HMI tags "Robot"
   "name" : Int, internal
   "DB1901_Config_Robots_Config_Robots{0}_Type_Kuka" : Bool = PLC DB1901_Config_Robots.Config_Robots[0].Type_Kuka AT %DB1901.DBX6.0, 1 s
      on ChangeValue: SetBit("DB1901_Config_Robots_Write")
   "DB1901_Config_Robots_Config_Robots{0}_Type_ABB" : Bool = PLC DB1901_Config_Robots.Config_Robots[0].Type_ABB AT %DB1901.DBX6.1, 1 s
      on ChangeValue: SetBit("DB1901_Config_Robots_Write")
   "DB1901_Config_Robots_Config_Robots{0}_Type_Fanuc" : Bool = PLC DB1901_Config_Robots.Config_Robots[0].Type_Fanuc AT %DB1901.DBX6.2, 1 s
      on ChangeValue: SetBit("DB1901_Config_Robots_Write")
   "DB1901_Config_Robots_Config_Robots{0}_Type_Motoman" : Bool = PLC DB1901_Config_Robots.Config_Robots[0].Type_Motoman AT %DB1901.DBX6.3, 1 s
      on ChangeValue: SetBit("DB1901_Config_Robots_Write")
   "DB1901_Config_Robots_Config_Robots{0}_Type_5" : Bool = PLC DB1901_Config_Robots.Config_Robots[0].Type_5 AT %DB1901.DBX6.4, 1 s
      on ChangeValue: SetBit("DB1901_Config_Robots_Write")
   "DB1901_Config_Robots_Config_Robots{0}_Type_6" : Bool = PLC DB1901_Config_Robots.Config_Robots[0].Type_6 AT %DB1901.DBX6.5, 1 s
      on ChangeValue: SetBit("DB1901_Config_Robots_Write")
   "DB1901_Config_Robots_Config_Robots{0}_Type_7" : Bool = PLC DB1901_Config_Robots.Config_Robots[0].Type_7 AT %DB1901.DBX6.6, 1 s
      on ChangeValue: SetBit("DB1901_Config_Robots_Write")
   "DB1901_Config_Robots_Config_Robots{0}_Type_8" : Bool = PLC DB1901_Config_Robots.Config_Robots[0].Type_8 AT %DB1901.DBX6.7, 1 s
      on ChangeValue: SetBit("DB1901_Config_Robots_Write")
   "DB1901_Config_Robots_Config_Robots{0}_With_Shotware" : Bool = PLC DB1901_Config_Robots.Config_Robots[0].With_Shotware AT %DB1901.DBX7.0, 1 s
      on ChangeValue: SetBit("DB1901_Config_Robots_Write")
   "DB1901_Config_Robots_Config_Robots{0}_With_Tracking" : Bool = PLC DB1901_Config_Robots.Config_Robots[0].With_Tracking AT %DB1901.DBX7.1, 1 s
      on ChangeValue: SetBit("DB1901_Config_Robots_Write")
   "DB1901_Config_Robots_Config_Robots{0}_With_Safetysoftware" : Bool = PLC DB1901_Config_Robots.Config_Robots[0].With_Safetysoftware AT %DB1901.DBX7.2, 1 s
      on ChangeValue: SetBit("DB1901_Config_Robots_Write")
   "DB1901_Config_Robots_Config_Robots{0}_With_Synchronisation" : Bool = PLC DB1901_Config_Robots.Config_Robots[0].With_Synchronisation AT %DB1901.DBX7.3, 1 s
      on ChangeValue: SetBit("DB1901_Config_Robots_Write")
   "DB1901_Config_Robots_Config_Robots{0}_With_Testshot" : Bool = PLC DB1901_Config_Robots.Config_Robots[0].With_Testshot AT %DB1901.DBX7.4, 1 s
      on ChangeValue: SetBit("DB1901_Config_Robots_Write")
   "DB1901_Config_Robots_Config_Robots{0}_With_Cleaning" : Bool = PLC DB1901_Config_Robots.Config_Robots[0].With_Cleaning AT %DB1901.DBX7.5, 1 s
      on ChangeValue: SetBit("DB1901_Config_Robots_Write")
   "DB1901_Config_Robots_Config_Robots{0}_With_Wet_Cleaning" : Bool = PLC DB1901_Config_Robots.Config_Robots[0].With_Wet_Cleaning AT %DB1901.DBX7.6, 1 s
      on ChangeValue: SetBit("DB1901_Config_Robots_Write")
   "DB1901_Config_Robots_Config_Robots{0}_With_Wet_Cleaning_LFI" : Bool = PLC DB1901_Config_Robots.Config_Robots[0].With_Wet_Cleaning_LFI AT %DB1901.DBX7.7, 1 s
      on ChangeValue: SetBit("DB1901_Config_Robots_Write")
   "DB1901_Config_Robots_Config_Robots{0}_With_Wet_Cleaning_Spray" : Bool = PLC DB1901_Config_Robots.Config_Robots[0].With_Wet_Cleaning_Spray AT %DB1901.DBX8.0, 1 s
      on ChangeValue: SetBit("DB1901_Config_Robots_Write")
   "DB1901_Config_Robots_Config_Robots{0}_With_IR_Station" : Bool = PLC DB1901_Config_Robots.Config_Robots[0].With_IR_Station AT %DB1901.DBX8.1, 1 s
      on ChangeValue: SetBit("DB1901_Config_Robots_Write")
   "DB1901_Config_Robots_Config_Robots{0}_With_Brush_Station" : Bool = PLC DB1901_Config_Robots.Config_Robots[0].With_Brush_Station AT %DB1901.DBX8.2, 1 s
      on ChangeValue: SetBit("DB1901_Config_Robots_Write")
   "DB1901_Config_Robots_Config_Robots{0}_With_Belt_Filter" : Bool = PLC DB1901_Config_Robots.Config_Robots[0].With_Belt_Filter AT %DB1901.DBX8.3, 1 s
      on ChangeValue: SetBit("DB1901_Config_Robots_Write")
   "DB1901_Config_Robots_Config_Robots{0}_With_Air_Cleaner" : Bool = PLC DB1901_Config_Robots.Config_Robots[0].With_Air_Cleaner AT %DB1901.DBX8.4, 1 s
      on ChangeValue: SetBit("DB1901_Config_Robots_Write")
   "DB1901_Config_Robots_Config_Robots{0}_Spare_2_5" : Bool = PLC DB1901_Config_Robots.Config_Robots[0].Spare_2_5 AT %DB1901.DBX8.5, 1 s
      on ChangeValue: SetBit("DB1901_Config_Robots_Write")
   "DB1901_Config_Robots_Config_Robots{0}_Spare_2_6" : Bool = PLC DB1901_Config_Robots.Config_Robots[0].Spare_2_6 AT %DB1901.DBX8.6, 1 s
      on ChangeValue: SetBit("DB1901_Config_Robots_Write")
   "DB1901_Config_Robots_Config_Robots{0}_Spare_2_7" : Bool = PLC DB1901_Config_Robots.Config_Robots[0].Spare_2_7 AT %DB1901.DBX8.7, 1 s
      on ChangeValue: SetBit("DB1901_Config_Robots_Write")
   "DB1900_IF_Robots_State_Robots{0}_EmergencyStopReady" : Bool = PLC DB1900_IF_Robots.State_Robots[0].EmergencyStopReady AT %DB1900.DBX96.4, 1 s
   "DB1900_IF_Robots_State_Robots{0}_AutomatcStopReady" : Bool = PLC DB1900_IF_Robots.State_Robots[0].AutomatcStopReady AT %DB1900.DBX96.5, 1 s
   "DB1900_IF_Robots_State_Robots{0}_MixingheadAuto" : Bool = PLC DB1900_IF_Robots.State_Robots[0].MixingheadAuto AT %DB1900.DBX96.6, 1 s
   "DB1900_IF_Robots_State_Robots{0}_MaschineAuto" : Bool = PLC DB1900_IF_Robots.State_Robots[0].MaschineAuto AT %DB1900.DBX96.7, 1 s
   "DB1900_IF_Robots_State_Robots{0}_TestShotRunning" : Bool = PLC DB1900_IF_Robots.State_Robots[0].TestShotRunning AT %DB1900.DBX97.3, 1 s
   "DB1900_IF_Robots_State_Robots{0}_Rob_in_Home" : Bool = PLC DB1900_IF_Robots.State_Robots[0].Rob_in_Home AT %DB1900.DBX96.0, 1 s
   "DB1900_IF_Robots_State_Robots{0}_Rob_in_Automatic" : Bool = PLC DB1900_IF_Robots.State_Robots[0].Rob_in_Automatic AT %DB1900.DBX96.1, 1 s
   "DB1900_IF_Robots_State_Robots{0}_Rob_in_Cycle" : Bool = PLC DB1900_IF_Robots.State_Robots[0].Rob_in_Cycle AT %DB1900.DBX96.2, 1 s
   "DB1900_IF_Robots_Switch_Robots{0}_SwitchHomePosON_OFF" : Bool = PLC DB1900_IF_Robots.Switch_Robots[0].SwitchHomePosON_OFF AT %DB1900.DBX6.0, 1 s
      on ChangeValue: SetBit("DB1900_IF_Robots_Write")
   "DB1900_IF_Robots_Switch_Robots{0}_SwitchMaintPosON_OFF" : Bool = PLC DB1900_IF_Robots.Switch_Robots[0].SwitchMaintPosON_OFF AT %DB1900.DBX6.1, 1 s
      on ChangeValue: SetBit("DB1900_IF_Robots_Write")
   "DB1900_IF_Robots_Switch_Robots{0}_SwitchMaintPos_2ON_OFF" : Bool = PLC DB1900_IF_Robots.Switch_Robots[0].SwitchMaintPos_2ON_OFF AT %DB1900.DBX6.2, 1 s
      on ChangeValue: SetBit("DB1900_IF_Robots_Write")
   "DB1900_IF_Robots_Switch_Robots{0}_SwitchTestShotON_OFF" : Bool = PLC DB1900_IF_Robots.Switch_Robots[0].SwitchTestShotON_OFF AT %DB1900.DBX6.3, 1 s
      on ChangeValue: SetBit("DB1900_IF_Robots_Write")
   "DB1900_IF_Robots_Switch_Robots{0}_SwitchCleaningON_OFF" : Bool = PLC DB1900_IF_Robots.Switch_Robots[0].SwitchCleaningON_OFF AT %DB1900.DBX6.4, 1 s
      on ChangeValue: SetBit("DB1900_IF_Robots_Write")
   "DB1900_IF_Robots_Switch_Robots{0}_SwitchBrushON_OFF" : Bool = PLC DB1900_IF_Robots.Switch_Robots[0].SwitchBrushON_OFF AT %DB1900.DBX6.5, 1 s
      on ChangeValue: SetBit("DB1900_IF_Robots_Write")
   "DB1900_IF_Robots_Switch_Robots{0}_SwitchSyncON_OFF" : Bool = PLC DB1900_IF_Robots.Switch_Robots[0].SwitchSyncON_OFF AT %DB1900.DBX6.6, 1 s
      on ChangeValue: SetBit("DB1900_IF_Robots_Write")
   "DB1900_IF_Robots_Switch_Robots{0}_SwitchTeachenON_OFF" : Bool = PLC DB1900_IF_Robots.Switch_Robots[0].SwitchTeachenON_OFF AT %DB1900.DBX6.7, 1 s
      on ChangeValue: SetBit("DB1900_IF_Robots_Write")
   "DB1900_IF_Robots_Switch_Robots{0}_SwitchLearningON_OFF" : Bool = PLC DB1900_IF_Robots.Switch_Robots[0].SwitchLearningON_OFF AT %DB1900.DBX7.0, 1 s
      on ChangeValue: SetBit("DB1900_IF_Robots_Write")
   "DB1900_IF_Robots_Switch_Robots{0}_SwitchAirCleaningON_OFF" : Bool = PLC DB1900_IF_Robots.Switch_Robots[0].SwitchAirCleaningON_OFF AT %DB1900.DBX7.1, 1 s
      on ChangeValue: SetBit("DB1900_IF_Robots_Write")
   "DB1900_IF_Robots_Switch_Robots{0}_SwitchAirCleaningManON_OFF" : Bool = PLC DB1900_IF_Robots.Switch_Robots[0].SwitchAirCleaningManON_OFF AT %DB1900.DBX7.2, 1 s
      on ChangeValue: SetBit("DB1900_IF_Robots_Write")
   "DB1900_IF_Robots_Switch_Robots{0}_StateHomePos" : Byte = PLC DB1900_IF_Robots.Switch_Robots[0].StateHomePos AT %DB1900.DBB8, 1 s
      on ChangeValue: SetBit("DB1900_IF_Robots_Write")
   "DB1900_IF_Robots_Switch_Robots{0}_StateMaintPos" : Byte = PLC DB1900_IF_Robots.Switch_Robots[0].StateMaintPos AT %DB1900.DBB9, 1 s
      on ChangeValue: SetBit("DB1900_IF_Robots_Write")
   "DB1900_IF_Robots_Switch_Robots{0}_StateMaintPos_2" : Byte = PLC DB1900_IF_Robots.Switch_Robots[0].StateMaintPos_2 AT %DB1900.DBB10, 1 s
      on ChangeValue: SetBit("DB1900_IF_Robots_Write")
   "DB1900_IF_Robots_Switch_Robots{0}_StateTestShot" : Byte = PLC DB1900_IF_Robots.Switch_Robots[0].StateTestShot AT %DB1900.DBB11, 1 s
      on ChangeValue: SetBit("DB1900_IF_Robots_Write")
   "DB1900_IF_Robots_Switch_Robots{0}_StateCleaning" : Byte = PLC DB1900_IF_Robots.Switch_Robots[0].StateCleaning AT %DB1900.DBB12, 1 s
      on ChangeValue: SetBit("DB1900_IF_Robots_Write")
   "DB1900_IF_Robots_Switch_Robots{0}_StateBrush" : Byte = PLC DB1900_IF_Robots.Switch_Robots[0].StateBrush AT %DB1900.DBB13, 1 s
      on ChangeValue: SetBit("DB1900_IF_Robots_Write")
   "DB1900_IF_Robots_Switch_Robots{0}_StateSync" : Byte = PLC DB1900_IF_Robots.Switch_Robots[0].StateSync AT %DB1900.DBB14, 1 s
      on ChangeValue: SetBit("DB1900_IF_Robots_Write")
   "DB1900_IF_Robots_Switch_Robots{0}_StateTeachen" : Byte = PLC DB1900_IF_Robots.Switch_Robots[0].StateTeachen AT %DB1900.DBB15, 1 s
      on ChangeValue: SetBit("DB1900_IF_Robots_Write")
   "DB1900_IF_Robots_Switch_Robots{0}_StateLearning" : Byte = PLC DB1900_IF_Robots.Switch_Robots[0].StateLearning AT %DB1900.DBB16, 1 s
      on ChangeValue: SetBit("DB1900_IF_Robots_Write")
   "DB1900_IF_Robots_Switch_Robots{0}_StateAirCleaning" : Byte = PLC DB1900_IF_Robots.Switch_Robots[0].StateAirCleaning AT %DB1900.DBB17, 1 s
      on ChangeValue: SetBit("DB1900_IF_Robots_Write")
   "DB1900_IF_Robots_Switch_Robots{0}_StateAirCleaningManual" : Byte = PLC DB1900_IF_Robots.Switch_Robots[0].StateAirCleaningManual AT %DB1900.DBB18, 1 s
      on ChangeValue: SetBit("DB1900_IF_Robots_Write")
   "DB1900_IF_Robots_ReadWriteDeviceNo" : Int = PLC DB1900_IF_Robots.ReadWriteDeviceNo AT %DB1900.DBW0, 1 s
   "DB1900_IF_Robots_Read" : Bool = PLC DB1900_IF_Robots.Read AT %DB1900.DBX4.0, 1 s
   "DB1900_IF_Robots_Write" : Bool = PLC DB1900_IF_Robots.Write AT %DB1900.DBX4.1, 1 s
   "DB1901_Config_Robots_Read" : Bool = PLC DB1901_Config_Robots.Read AT %DB1901.DBX4.0, 1 s
   "DB1901_Config_Robots_Write" : Bool = PLC DB1901_Config_Robots.Write AT %DB1901.DBX4.1, 1 s
   "DB1900_IF_Robots_State_Robots{0}_Rob_Prog_No" : Byte = PLC DB1900_IF_Robots.State_Robots[0].Rob_Prog_No AT %DB1900.DBB98, 1 s
   "DB1900_IF_Robots_State_Robots{0}_Rob_MC_No" : Byte = PLC DB1900_IF_Robots.State_Robots[0].Rob_MC_No AT %DB1900.DBB99, 1 s

HMI tags "Navigation Button"
   "DB14_TP_Shortcuts_TP_Shortcuts_ButtonNo_1" : Bool = PLC DB14_TP_Shortcuts.TP_Shortcuts.ButtonNo.1, 1 s
   "DB14_TP_Shortcuts_TP_Shortcuts_ButtonNo_2" : Bool = PLC DB14_TP_Shortcuts.TP_Shortcuts.ButtonNo.2, 1 s
   "DB14_TP_Shortcuts_TP_Shortcuts_ButtonNo_3" : Bool = PLC DB14_TP_Shortcuts.TP_Shortcuts.ButtonNo.3, 1 s
   "DB14_TP_Shortcuts_TP_Shortcuts_ButtonNo_5" : Bool = PLC DB14_TP_Shortcuts.TP_Shortcuts.ButtonNo.5, 1 s
   "DB14_TP_Shortcuts_TP_Shortcuts_ButtonNo_6" : Bool = PLC DB14_TP_Shortcuts.TP_Shortcuts.ButtonNo.6, 1 s
   "DB14_TP_Shortcuts_TP_Shortcuts_ButtonNo_7" : Bool = PLC DB14_TP_Shortcuts.TP_Shortcuts.ButtonNo.7, 1 s
   "DB14_TP_Shortcuts_TP_Shortcuts_Page_active_1" : Bool = PLC DB14_TP_Shortcuts.TP_Shortcuts.Page_active.1, 1 s
   "DB14_TP_Shortcuts_TP_Shortcuts_Page_active_2" : Bool = PLC DB14_TP_Shortcuts.TP_Shortcuts.Page_active.2, 1 s
   "DB14_TP_Shortcuts_TP_Shortcuts_Page_active_3" : Bool = PLC DB14_TP_Shortcuts.TP_Shortcuts.Page_active.3, 1 s
   "DB14_TP_Shortcuts_TP_Shortcuts_Page_active_4" : Bool = PLC DB14_TP_Shortcuts.TP_Shortcuts.Page_active.4, 1 s
   "DB14_TP_Shortcuts_TP_Shortcuts_Page_active_5" : Bool = PLC DB14_TP_Shortcuts.TP_Shortcuts.Page_active.5, 1 s
   "DB14_TP_Shortcuts_TP_Shortcuts_Page_active_6" : Bool = PLC DB14_TP_Shortcuts.TP_Shortcuts.Page_active.6, 1 s
   "DB14_TP_Shortcuts_TP_Shortcuts_Page_active_7" : Bool = PLC DB14_TP_Shortcuts.TP_Shortcuts.Page_active.7, 1 s
   "DB14_TP_Shortcuts_TP_Shortcuts_PageNo_1" : Int = PLC DB14_TP_Shortcuts.TP_Shortcuts.PageNo.1, 1 s
   "DB14_TP_Shortcuts_TP_Shortcuts_PageNo_2" : Int = PLC DB14_TP_Shortcuts.TP_Shortcuts.PageNo.2, 1 s
   "DB14_TP_Shortcuts_TP_Shortcuts_PageNo_3" : Int = PLC DB14_TP_Shortcuts.TP_Shortcuts.PageNo.3, 1 s
   "DB14_TP_Shortcuts_TP_Shortcuts_PageNo_4" : Int = PLC DB14_TP_Shortcuts.TP_Shortcuts.PageNo.4, 1 s
   "DB14_TP_Shortcuts_TP_Shortcuts_PageNo_5" : Int = PLC DB14_TP_Shortcuts.TP_Shortcuts.PageNo.5, 1 s
   "DB14_TP_Shortcuts_TP_Shortcuts_PageNo_6" : Int = PLC DB14_TP_Shortcuts.TP_Shortcuts.PageNo.6, 1 s
   "DB14_TP_Shortcuts_TP_Shortcuts_PageNo_7" : Int = PLC DB14_TP_Shortcuts.TP_Shortcuts.PageNo.7, 1 s
   "Navigation_7" : Int, internal

discrete alarms
   1: 'Machine 01: Data loss after control general reset', class Machine Alarm Warning, trigger "Machine_Alarm_DBW_58" bit 8
   2: 'Machine 01: Fuse Fault', class Machine Alarm Warning, trigger "Machine_Alarm_DBW_58" bit 9
   3: 'Machine 01: Connection to computer faultly', class Machine Alarm Warning, trigger "Machine_Alarm_DBW_58" bit 10
   4: 'Machine 01: Control Cabinet Door Open', class Machine Alarm Warning, trigger "Machine_Alarm_DBW_58" bit 11
   5: 'Machine 01: Air Drier fault', class Machine Alarm Warning, trigger "Machine_Alarm_DBW_58" bit 12
   6: 'Machine 01: Control Voltage missing', class Machine Warning Archive Foaming, trigger "Machine_Alarm_DBW_58" bit 13
   7: 'Machine 01: Plunger Service not permitted', class Machine Alarm Warning, trigger "Machine_Alarm_DBW_58" bit 14
   8: 'Machine 01: Fuse fault on mixinghead', class Machine Alarm Warning, trigger "Machine_Alarm_DBW_58" bit 15
   9: 'Machine 01: Heater fault', class Machine Alarm Warning, trigger "Machine_Alarm_DBW_58" bit 0
   10: 'Machine 01: IMM fault', class Machine Alarm Warning, trigger "Machine_Alarm_DBW_58" bit 1
   11: 'Machine 01: Fuse fault on cooler', class Machine Alarm Warning, trigger "Machine_Alarm_DBW_58" bit 2
   12: 'Machine 01: Incorrect mix.ing head number', class Machine Alarm Warning, trigger "Machine_Alarm_DBW_58" bit 3
   13: 'Machine 01: Fuse fault, plasma', class Machine Alarm Warning, trigger "Machine_Alarm_DBW_58" bit 4
   14: 'Machine 01: Run empty day tank is selected', class Machine Alarm Warning, trigger "Machine_Alarm_DBW_58" bit 5
   15: 'Machine 01: IMM not in automatic', class Machine Alarm Warning, trigger "Machine_Alarm_DBW_58" bit 6
   16: 'Machine 01: Spare', class Machine Alarm Warning, trigger "Machine_Alarm_DBW_58" bit 7
   17: 'Machine 01: Machine emergency stop actuated', class Machine Warning Archive Foaming, trigger "Machine_Alarm_DBW_60" bit 8
   18: 'Machine 01: Emergency stop actuated at the control cabinet', class Machine Alarm Warning, trigger "Machine_Alarm_DBW_60" bit 9
   19: 'Machine 01: Emergency stop actuated at the control panel', class Machine Alarm Warning, trigger "Machine_Alarm_DBW_60" bit 10
   20: 'Machine 01: Emergency stop actuated at second monitor', class Machine Alarm Warning, trigger "Machine_Alarm_DBW_60" bit 11
   21: 'Machine 01: Emergency stop actuated at day tank', class Machine Alarm Warning, trigger "Machine_Alarm_DBW_60" bit 12
   22: 'Machine 01: Emergency stop actuated at the mixinghead clean', class Machine Alarm Warning, trigger "Machine_Alarm_DBW_60" bit 13
   23: 'Machine 01: Emergency stop actuated at nucleation unit', class Machine Alarm Warning, trigger "Machine_Alarm_DBW_60" bit 14
   24: 'Machine 01: Robot emergency stop pending', class Machine Alarm Warning, trigger "Machine_Alarm_DBW_60" bit 15
   25: 'Machine 01: Robot 2 emergency stop pending', class Machine Alarm Warning, trigger "Machine_Alarm_DBW_60" bit 0
   26: 'Machine 01: Container station emer. stop pending', class Machine Alarm Warning, trigger "Machine_Alarm_DBW_60" bit 1
   27: 'Machine 01: Container 2 emergency stop pending', class Machine Alarm Warning, trigger "Machine_Alarm_DBW_60" bit 2
   28: 'Machine 01: Emergency stop external system pending', class Machine Alarm Warning, trigger "Machine_Alarm_DBW_60" bit 3
   29: 'Machine 01: Emergency stop external system pending', class Machine Alarm Warning, trigger "Machine_Alarm_DBW_60" bit 4
   30: 'Machine 01: Emergency stop colour metering pending', class Machine Alarm Warning, trigger "Machine_Alarm_DBW_60" bit 5
   31: 'Machine 01: Emergency stop colour metering 2 pending', class Machine Alarm Warning, trigger "Machine_Alarm_DBW_60" bit 6
   32: 'Machine 01: Emergency stop from a mould carrier pending', class Machine Alarm Warning, trigger "Machine_Alarm_DBW_60" bit 7
   33: 'Machine 01: Operation mode test is selected', class Machine Warning Archive Foaming, trigger "Machine_Alarm_DBW_62" bit 8
   34: 'Machine 01: Weekend mode is activated', class Machine Alarm Warning, trigger "Machine_Alarm_DBW_62" bit 9
   35: 'Machine 01: Interface PC', class Machine Alarm Warning, trigger "Machine_Alarm_DBW_62" bit 10
   36: 'Machine 01: Buffer batery fault', class Machine Alarm Warning, trigger "Machine_Alarm_DBW_62" bit 11
   37: 'Machine 01: Automatic stop still not acknowledged', class Machine Alarm Warning, trigger "Machine_Alarm_DBW_62" bit 12
   38: 'Machine 01: Fault, pentane pre-alarm', class Machine Alarm Warning, trigger "Machine_Alarm_DBW_62" bit 13
   39: 'Machine 01: Fault, pentane alarm', class Machine Alarm Warning, trigger "Machine_Alarm_DBW_62" bit 14
   40: 'Machine 01: Air supply fault', class Machine Alarm Warning, trigger "Machine_Alarm_DBW_62" bit 15
   41: 'Machine 01: Computer fault group 1', class Machine Alarm Warning, trigger "Machine_Alarm_DBW_62" bit 0
   42: 'Machine 01: Computer fault group 2', class Machine Alarm Warning, trigger "Machine_Alarm_DBW_62" bit 1
   43: 'Machine 01: Computer fault group 3', class Machine Alarm Warning, trigger "Machine_Alarm_DBW_62" bit 2
   44: 'Machine 01: Spare', class Machine Alarm Warning, trigger "Machine_Alarm_DBW_62" bit 3
   45: 'Machine 01: Data buffer for foaming data is full!', class Machine Alarm Warning, trigger "Machine_Alarm_DBW_62" bit 4
   46: 'Machine 01: Error when writing to MMC', class Machine Alarm Warning, trigger "Machine_Alarm_DBW_62" bit 5
   47: 'Machine 01: Watchdog', class Machine Alarm Warning, trigger "Machine_Alarm_DBW_62" bit 6
   48: 'Machine 01: Container station not ready', class Machine Alarm Warning, trigger "Machine_Alarm_DBW_62" bit 7
   49: 'Machine 01: Shot time is too short', class Machine Alarm Warning, trigger "Machine_Alarm_DBW_64" bit 8
   50: 'Machine 01: Tool cannot be removed', class Machine Alarm Warning, trigger "Machine_Alarm_DBW_64" bit 9
   51: 'Machine 01: Pneumatic-pressure at supply is not available', class Machine Alarm Warning, trigger "Machine_Alarm_DBW_64" bit 10
   52: 'Machine 01: Pneumatic -pressure at smooth start is not available', class Machine Alarm Warning, trigger "Machine_Alarm_DBW_64" bit 11
   53: 'Machine 01: Spare', class Machine Alarm Warning, trigger "Machine_Alarm_DBW_64" bit 12
   54: 'Machine 01: Spare', class Machine Alarm Warning, trigger "Machine_Alarm_DBW_64" bit 13
   55: 'Machine 01: Spare', class Machine Alarm Warning, trigger "Machine_Alarm_DBW_64" bit 14
   56: 'Machine 01: Spare', class Machine Alarm Warning, trigger "Machine_Alarm_DBW_64" bit 15
   57: 'Machine 01: Time value for runtime or pause time incorrect', class Machine Alarm Warning, trigger "Machine_Alarm_DBW_64" bit 0
   58: 'Machine 01:', class Machine Alarm Warning, trigger "Machine_Alarm_DBW_64" bit 1
   59: 'Machine 01:', class Machine Alarm Warning, trigger "Machine_Alarm_DBW_64" bit 2
   60: 'Machine 01:', class Machine Alarm Warning, trigger "Machine_Alarm_DBW_64" bit 3
   61: 'Machine 01:', class Machine Alarm Warning, trigger "Machine_Alarm_DBW_64" bit 4
   62: 'Machine 01:', class Machine Alarm Warning, trigger "Machine_Alarm_DBW_64" bit 5
   63: 'Machine 01:', class Machine Alarm Warning, trigger "Machine_Alarm_DBW_64" bit 6
   64: 'Machine 01:', class Machine Alarm Warning, trigger "Machine_Alarm_DBW_64" bit 7
   501: 'General: fault Profinet: ProNet Module 01', class Machine Warning Archive Foaming, trigger "Profibus_Alarm_DBW_16" bit 8
   502: 'General: fault Profinet: ProNet Module 02', class Machine Warning Archive Foaming, trigger "Profibus_Alarm_DBW_16" bit 9
   503: 'General: fault Profinet: pn-pn coupler', class Machine Warning Archive Foaming, trigger "Profibus_Alarm_DBW_16" bit 10
   504: 'General: fault Profibus user 04', class Machine Alarm Warning, trigger "Profibus_Alarm_DBW_16" bit 11
   505: 'General: fault Profibus user 05', class Machine Alarm Warning, trigger "Profibus_Alarm_DBW_16" bit 12
   506: 'General: fault Profibus user 06', class Machine Alarm Warning, trigger "Profibus_Alarm_DBW_16" bit 13
   507: 'General: fault Profibus user 07', class Machine Alarm Warning, trigger "Profibus_Alarm_DBW_16" bit 14
   508: 'General: fault Profibus user 08', class Machine Alarm Warning, trigger "Profibus_Alarm_DBW_16" bit 15
   509: 'General: fault Profibus user 09', class Machine Alarm Warning, trigger "Profibus_Alarm_DBW_16" bit 0
   510: 'General: fault Profibus user 10', class Machine Alarm Warning, trigger "Profibus_Alarm_DBW_16" bit 1
   511: 'General: fault Profibus user 11 // ProCan module in terminal box for mixing head', class Machine Alarm Warning, trigger "Profibus_Alarm_DBW_16" bit 2
   512: 'General: fault Profibus user 12', class Machine Alarm Warning, trigger "Profibus_Alarm_DBW_16" bit 3
   513: 'General: fault Profibus user 13', class Machine Alarm Warning, trigger "Profibus_Alarm_DBW_16" bit 4
   514: 'General: fault Profibus user 14', class Machine Alarm Warning, trigger "Profibus_Alarm_DBW_16" bit 5
   515: 'General: fault Profibus user 15 //DP//DP Coupler', class Machine Alarm Warning, trigger "Profibus_Alarm_DBW_16" bit 6
   516: 'General: fault Profibus user 16', class Machine Alarm Warning, trigger "Profibus_Alarm_DBW_16" bit 7
   517: 'General: fault Profibus user 17', class Machine Alarm Warning, trigger "Profibus_Alarm_DBW_18" bit 8
   518: 'General: fault Profibus user 18', class Machine Alarm Warning, trigger "Profibus_Alarm_DBW_18" bit 9
   519: 'General: fault Profibus user 19', class Machine Alarm Warning, trigger "Profibus_Alarm_DBW_18" bit 10
   520: 'General: fault Profibus user 20', class Machine Alarm Warning, trigger "Profibus_Alarm_DBW_18" bit 11
   521: 'General: fault Profibus user 21 // ProCan module in terminal box for mixing head', class Machine Alarm Warning, trigger "Profibus_Alarm_DBW_18" bit 12
   522: 'General:', class Machine Alarm Warning, trigger "Profibus_Alarm_DBW_18" bit 13
   523: 'General:', class Machine Alarm Warning, trigger "Profibus_Alarm_DBW_18" bit 14
   524: 'General:', class Machine Alarm Warning, trigger "Profibus_Alarm_DBW_18" bit 15
   525: 'General:', class Machine Alarm Warning, trigger "Profibus_Alarm_DBW_18" bit 0
   526: 'General:', class Machine Alarm Warning, trigger "Profibus_Alarm_DBW_18" bit 1
   527: 'General:', class Machine Alarm Warning, trigger "Profibus_Alarm_DBW_18" bit 2
   528: 'General:', class Machine Alarm Warning, trigger "Profibus_Alarm_DBW_18" bit 3
   529: 'General:', class Machine Alarm Warning, trigger "Profibus_Alarm_DBW_18" bit 4
   530: 'General:', class Machine Alarm Warning, trigger "Profibus_Alarm_DBW_18" bit 5
   531: 'General: fault Profibus user 31 // ProCan module in terminal box for mixing head', class Machine Alarm Warning, trigger "Profibus_Alarm_DBW_18" bit 6
   532: 'General:', class Machine Alarm Warning, trigger "Profibus_Alarm_DBW_18" bit 7
   533: 'General:', class Machine Alarm Warning, trigger "Profibus_Alarm_DBW_20" bit 8
   534: 'General:', class Machine Alarm Warning, trigger "Profibus_Alarm_DBW_20" bit 9
   535: 'General:', class Machine Alarm Warning, trigger "Profibus_Alarm_DBW_20" bit 10
   536: 'General:', class Machine Alarm Warning, trigger "Profibus_Alarm_DBW_20" bit 11
   537: 'General:', class Machine Alarm Warning, trigger "Profibus_Alarm_DBW_20" bit 12
   538: 'General:', class Machine Alarm Warning, trigger "Profibus_Alarm_DBW_20" bit 13
   539: 'General:', class Machine Alarm Warning, trigger "Profibus_Alarm_DBW_20" bit 14
   540: 'General:', class Machine Alarm Warning, trigger "Profibus_Alarm_DBW_20" bit 15
   541: 'General: fault Profibus user 41 // ProCan module in terminal box for mixing head', class Machine Alarm Warning, trigger "Profibus_Alarm_DBW_20" bit 0
   542: 'General:', class Machine Alarm Warning, trigger "Profibus_Alarm_DBW_20" bit 1
   543: 'General:', class Machine Alarm Warning, trigger "Profibus_Alarm_DBW_20" bit 2
   544: 'General:', class Machine Alarm Warning, trigger "Profibus_Alarm_DBW_20" bit 3
   545: 'General:', class Machine Alarm Warning, trigger "Profibus_Alarm_DBW_20" bit 4
   546: 'General:', class Machine Alarm Warning, trigger "Profibus_Alarm_DBW_20" bit 5
   547: 'General:', class Machine Alarm Warning, trigger "Profibus_Alarm_DBW_20" bit 6
   548: 'General:', class Machine Alarm Warning, trigger "Profibus_Alarm_DBW_20" bit 7
   549: 'General:', class Machine Alarm Warning, trigger "Profibus_Alarm_DBW_22" bit 8
   550: 'General:', class Machine Alarm Warning, trigger "Profibus_Alarm_DBW_22" bit 9
   551: 'General: fault Profibus user 51 // ProCan module in terminal box for mixing head', class Machine Alarm Warning, trigger "Profibus_Alarm_DBW_22" bit 10
   552: 'General:', class Machine Alarm Warning, trigger "Profibus_Alarm_DBW_22" bit 11
   553: 'General:', class Machine Alarm Warning, trigger "Profibus_Alarm_DBW_22" bit 12
   554: 'General:', class Machine Alarm Warning, trigger "Profibus_Alarm_DBW_22" bit 13
   555: 'General:', class Machine Alarm Warning, trigger "Profibus_Alarm_DBW_22" bit 14
   556: 'General:', class Machine Alarm Warning, trigger "Profibus_Alarm_DBW_22" bit 15
   565: 'General:', class Machine Alarm Warning, trigger "Profibus_Alarm_DBW_24" bit 8
   566: 'General:', class Machine Alarm Warning, trigger "Profibus_Alarm_DBW_24" bit 9
   567: 'General:', class Machine Alarm Warning, trigger "Profibus_Alarm_DBW_24" bit 10
   568: 'General:', class Machine Alarm Warning, trigger "Profibus_Alarm_DBW_24" bit 11
   569: 'General:', class Machine Alarm Warning, trigger "Profibus_Alarm_DBW_24" bit 12
   570: 'General:', class Machine Alarm Warning, trigger "Profibus_Alarm_DBW_24" bit 13
   571: 'General: fault Profibus user 71 // ProCan module in terminal box for mixing head', class Machine Alarm Warning, trigger "Profibus_Alarm_DBW_24" bit 14
   572: 'General:', class Machine Alarm Warning, trigger "Profibus_Alarm_DBW_24" bit 15
   573: 'General:', class Machine Alarm Warning, trigger "Profibus_Alarm_DBW_24" bit 0
   574: 'General:', class Machine Alarm Warning, trigger "Profibus_Alarm_DBW_24" bit 1
   575: 'General:', class Machine Alarm Warning, trigger "Profibus_Alarm_DBW_24" bit 2
   576: 'General:', class Machine Alarm Warning, trigger "Profibus_Alarm_DBW_24" bit 3
   577: 'General:', class Machine Alarm Warning, trigger "Profibus_Alarm_DBW_24" bit 4
   578: 'General:', class Machine Alarm Warning, trigger "Profibus_Alarm_DBW_24" bit 5
   579: 'General:', class Machine Alarm Warning, trigger "Profibus_Alarm_DBW_24" bit 6
   580: 'General:', class Machine Alarm Warning, trigger "Profibus_Alarm_DBW_24" bit 7
   581: 'General: fault Profibus user 81 // ProCan module in terminal box for mixinghead', class Machine Alarm Warning, trigger "Profibus_Alarm_DBW_26" bit 8
   582: 'General:', class Machine Alarm Warning, trigger "Profibus_Alarm_DBW_26" bit 9
   583: 'General:', class Machine Alarm Warning, trigger "Profibus_Alarm_DBW_26" bit 10
   584: 'General:', class Machine Alarm Warning, trigger "Profibus_Alarm_DBW_26" bit 11
   585: 'General:', class Machine Alarm Warning, trigger "Profibus_Alarm_DBW_26" bit 12
   586: 'General:', class Machine Alarm Warning, trigger "Profibus_Alarm_DBW_26" bit 13
   587: 'General:', class Machine Alarm Warning, trigger "Profibus_Alarm_DBW_26" bit 14
   588: 'General:', class Machine Alarm Warning, trigger "Profibus_Alarm_DBW_26" bit 15
   589: 'General:', class Machine Alarm Warning, trigger "Profibus_Alarm_DBW_26" bit 0
   590: 'General:', class Machine Alarm Warning, trigger "Profibus_Alarm_DBW_26" bit 1
   591: 'General: fault Profibus user 91 // ProCan module in terminal box for mixing head', class Machine Alarm Warning, trigger "Profibus_Alarm_DBW_26" bit 2
   592: 'General:', class Machine Alarm Warning, trigger "Profibus_Alarm_DBW_26" bit 3
   593: 'General:', class Machine Alarm Warning, trigger "Profibus_Alarm_DBW_26" bit 4
   594: 'General:', class Machine Alarm Warning, trigger "Profibus_Alarm_DBW_26" bit 5
   595: 'General:', class Machine Alarm Warning, trigger "Profibus_Alarm_DBW_26" bit 6
   596: 'General:', class Machine Alarm Warning, trigger "Profibus_Alarm_DBW_26" bit 7
   597: 'General:', class Machine Alarm Warning, trigger "Profibus_Alarm_DBW_28" bit 8
   598: 'General:', class Machine Alarm Warning, trigger "Profibus_Alarm_DBW_28" bit 9
   599: 'General:', class Machine Alarm Warning, trigger "Profibus_Alarm_DBW_28" bit 10
   600: 'General: fault Profibus user 100', class Machine Alarm Warning, trigger "Profibus_Alarm_DBW_28" bit 11
   601: 'General: fault Profibus user 101 // ProCan Module in terminal box for mixinghead', class Machine Alarm Warning, trigger "Profibus_Alarm_DBW_28" bit 12
   557: 'Machine 01:', class Machine Alarm Warning, trigger "Profibus_Alarm_DBW_22" bit 0
   558: 'Machine 01:', class Machine Alarm Warning, trigger "Profibus_Alarm_DBW_22" bit 1
   559: 'Machine 01:', class Machine Alarm Warning, trigger "Profibus_Alarm_DBW_22" bit 2
   560: 'Machine 01:', class Machine Alarm Warning, trigger "Profibus_Alarm_DBW_22" bit 3
   561: 'Machine 01:', class Machine Alarm Warning, trigger "Profibus_Alarm_DBW_22" bit 4
   562: 'Machine 01:', class Machine Alarm Warning, trigger "Profibus_Alarm_DBW_22" bit 5
   563: 'Machine 01:', class Machine Alarm Warning, trigger "Profibus_Alarm_DBW_22" bit 6
   564: 'Machine 01:', class Machine Alarm Warning, trigger "Profibus_Alarm_DBW_22" bit 7
   602: 'Machine 01:', class Machine Alarm Warning, trigger "Profibus_Alarm_DBW_28" bit 13
   603: 'Machine 01:', class Machine Alarm Warning, trigger "Profibus_Alarm_DBW_28" bit 14
   604: 'Machine 01:', class Machine Alarm Warning, trigger "Profibus_Alarm_DBW_28" bit 15
   605: 'Machine 01:', class Machine Alarm Warning, trigger "Profibus_Alarm_DBW_28" bit 0
   701: 'TankTank1:', class Tank Alarm Warning, trigger "Interface_Container_DBW_520" bit 8
   702: 'TankTank1:', class Tank Alarm Warning, trigger "Interface_Container_DBW_520" bit 9
   703: 'TankTank1:', class Tank Alarm Warning, trigger "Interface_Container_DBW_520" bit 10
   704: 'TankTank1:', class Tank Alarm Warning, trigger "Interface_Container_DBW_520" bit 11
   705: 'ContainerStation: Station Tank1 not ready', class Tank Alarm Warning, trigger "Interface_Container_DBW_520" bit 12
   706: 'ContainerStation: Station Tank2 not ready', class Tank Alarm Warning, trigger "Interface_Container_DBW_520" bit 13
   707: 'TankTank1:', class Tank Alarm Warning, trigger "Interface_Container_DBW_520" bit 14
   708: 'TankTank1:', class Tank Alarm Warning, trigger "Interface_Container_DBW_520" bit 15
   709: 'TankTank1:', class Tank Alarm Warning, trigger "Interface_Container_DBW_520" bit 0
   710: 'TankTank1:', class Tank Alarm Warning, trigger "Interface_Container_DBW_520" bit 1
   711: 'TankTank1:', class Tank Alarm Warning, trigger "Interface_Container_DBW_520" bit 2
   712: 'TankTank1:', class Tank Alarm Warning, trigger "Interface_Container_DBW_520" bit 3
   11101: 'Tank Tank1: Feed Pump: Motor Protecting switch has tripped', class Tank Alarm Warning, trigger "Tank1_FeedPump_DBW_2" bit 8
   11102: 'Tank Tank1: Feed Pump: Frequency converter fault', class Tank Alarm Warning, trigger "Tank1_FeedPump_DBW_2" bit 9
   11103: 'Tank Tank1: Feed Pump: Max.Pressure', class Tank Alarm Warning, trigger "Tank1_FeedPump_DBW_2" bit 10
   11104: 'Tank Tank1: Feed Pump: Dry run protection has tripped', class Tank Alarm Warning, trigger "Tank1_FeedPump_DBW_2" bit 11
   11105: 'Tank Tank1: Feed Pump: Wrong time entry for pause and runtime', class Tank Alarm Warning, trigger "Tank1_FeedPump_DBW_2" bit 12
   11106: 'Tank Tank1: Feed Pump: Difference pressure too high', class Tank Alarm Warning, trigger "Tank1_FeedPump_DBW_2" bit 13
   11107: 'Tank Tank1: Feed Pump: Temperature for switch-on not reached', class Tank Alarm Warning, trigger "Tank1_FeedPump_DBW_2" bit 14
   11108: 'Tank Tank1: Feed Pump: Motor protecting switch fan has tripped', class Tank Alarm Warning, trigger "Tank1_FeedPump_DBW_2" bit 15
   11109: 'Tank Tank1: Feed Pump: Filling level too low', class Tank Alarm Warning, trigger "Tank1_FeedPump_DBW_2" bit 0
   11110: 'Tank Tank1: Feed Pump: Filling selected but no barrel present', class Tank Alarm Warning, trigger "Tank1_FeedPump_DBW_2" bit 1
   11111: 'Tank Tank1: Feed Pump: No barrel present', class Tank Caution, trigger "Tank1_FeedPump_DBW_2" bit 2
   11112: 'Tank Tank1: Feed Pump:', class Tank Alarm Warning, trigger "Tank1_FeedPump_DBW_2" bit 3
   11113: 'Tank Tank1: Feed Pump:', class Tank Alarm Warning, trigger "Tank1_FeedPump_DBW_2" bit 4
   11114: 'Tank Tank1: Feed Pump:', class Tank Alarm Warning, trigger "Tank1_FeedPump_DBW_2" bit 5
   11115: 'Tank Tank1: Feed Pump:', class Tank Alarm Warning, trigger "Tank1_FeedPump_DBW_2" bit 6
   11116: 'Tank Tank1: Feed Pump:', class Tank Alarm Warning, trigger "Tank1_FeedPump_DBW_2" bit 7
   11117: 'Tank Tank1: Agitator: Motor protecting switch has tripped', class Tank Alarm Warning, trigger "Tank1_Agitator_DBW_28" bit 8
   11118: 'Tank Tank1: Agitator: Frequencny converter fault', class Tank Alarm Warning, trigger "Tank1_Agitator_DBW_28" bit 9
   11119: 'Tank Tank1: Agitator: Max drip pan filling level', class Tank Alarm Warning, trigger "Tank1_Agitator_DBW_28" bit 10
   11120: 'Tank Tank1: Agitator: Incorrect time entry for runtime or pause time', class Tank Alarm Warning, trigger "Tank1_Agitator_DBW_28" bit 11
   11121: 'Tank Tank1: Agitator:', class Tank Alarm Warning, trigger "Tank1_Agitator_DBW_28" bit 12
   11122: 'Tank Tank1: Agitator: Temperature for switch-on not reached', class Tank Alarm Warning, trigger "Tank1_Agitator_DBW_28" bit 13
   11123: 'Tank Tank1: Agitator: Fan motor protecting switch', class Tank Alarm Warning, trigger "Tank1_Agitator_DBW_28" bit 14
   11124: 'Tank Tank1: Agitator: Filling level too low', class Tank Alarm Warning, trigger "Tank1_Agitator_DBW_28" bit 15
   11125: 'Tank Tank1: Agitator:', class Tank Alarm Warning, trigger "Tank1_Agitator_DBW_28" bit 0
   11126: 'Tank Tank1: Agitator:', class Tank Alarm Warning, trigger "Tank1_Agitator_DBW_28" bit 1
   11127: 'Tank Tank1: Agitator:', class Tank Alarm Warning, trigger "Tank1_Agitator_DBW_28" bit 2
   11128: 'Tank Tank1: Agitator:', class Tank Alarm Warning, trigger "Tank1_Agitator_DBW_28" bit 3
   11129: 'Tank Tank1: Agitator:', class Tank Alarm Warning, trigger "Tank1_Agitator_DBW_28" bit 4
   11130: 'Tank Tank1: Agitator:', class Tank Alarm Warning, trigger "Tank1_Agitator_DBW_28" bit 5
   11131: 'Tank Tank1: Agitator:', class Tank Alarm Warning, trigger "Tank1_Agitator_DBW_28" bit 6
   11133: 'Tank Tank1: Filling: Min. filling level undershot', class Tank Warning Archive Foaming, trigger "Tank1_Filling_DBW_54" bit 8
   11134: 'Tank Tank1: Filling: Max. filling level exceeded', class Tank Warning Archive Foaming, trigger "Tank1_Filling_DBW_54" bit 9
   11135: 'Tank Tank1: Filling: Filling time exceeded', class Tank Alarm Warning, trigger "Tank1_Filling_DBW_54" bit 10
   11136: 'Tank Tank1: Filling: Max. drip pan filling level', class Tank Alarm Warning, trigger "Tank1_Filling_DBW_54" bit 11
   11137: 'Tank Tank1: Filling: Min. filling level in cycle', class Tank Error Filling, trigger "Tank1_Filling_DBW_54" bit 12
   11138: 'Tank Tank1: Filling: Max. filling level (with piston machines)', class Tank Error, trigger "Tank1_Filling_DBW_54" bit 13
   11139: 'Tank Tank1: Filling: Max. drip pan filling level (with piston machines)', class Tank Error Filling, trigger "Tank1_Filling_DBW_54" bit 14
   11140: 'Tank Tank1: Filling: Cable break to fill level sensor', class Tank Error Filling, trigger "Tank1_Filling_DBW_54" bit 15
   11141: 'Tank Tank1: Filling: Wrong position of fill valve', class Tank Error Filling, trigger "Tank1_Filling_DBW_54" bit 0
   11142: 'Tank Tank1: Filling: Pre-warning min. filling level', class Tank Errors Fill Archive Foaming, trigger "Tank1_Filling_DBW_54" bit 1
   11143: 'Tank Tank1: Filling:', class Tank Error Filling, trigger "Tank1_Filling_DBW_54" bit 2
   11144: 'Tank Tank1: Filling:', class Tank Error Filling, trigger "Tank1_Filling_DBW_54" bit 3
   11145: 'Tank Tank1: Filling:', class Tank Error Filling, trigger "Tank1_Filling_DBW_54" bit 4
   11146: 'Tank Tank1: Filling: Motor protection supply nucleation unit', class Tank Error Filling, trigger "Tank1_Filling_DBW_54" bit 5
   11147: 'Tank Tank1: Filling: Cable break analog value of nucleation unit', class Tank Error Filling, trigger "Tank1_Filling_DBW_54" bit 6
   11148: 'Tank Tank1: Filling: Fault from nucleation unit', class Tank Error Filling, trigger "Tank1_Filling_DBW_54" bit 7
   11149: 'Tank Tank1: Heat-balancing: Cable break to temperature sensor', class Tank Errors Archive Foaming, trigger "Tank1_ControlerTemp_DBW_236" bit 8
   11150: 'Tank Tank1: Heat-balancing: + Temperature warning', class Tank Alarm Warning, trigger "Tank1_ControlerTemp_DBW_236" bit 9
   11151: 'Tank Tank1: Heat-balancing: - Temperature warning', class Tank Alarm Warning, trigger "Tank1_ControlerTemp_DBW_236" bit 10
   11152: 'Tank Tank1: Heat-balancing: + Temperature fault', class Tank Error, trigger "Tank1_ControlerTemp_DBW_236" bit 11
   11153: 'Tank Tank1: Heat-balancing: - Temperature fault', class Tank Error, trigger "Tank1_ControlerTemp_DBW_236" bit 12
   11154: 'Tank Tank1: Heat-balancing:Controller at limit', class Tank Alarm Warning, trigger "Tank1_ControlerTemp_DBW_236" bit 13
   11155: 'Tank Tank1: Heat-balancing:', class Tank Alarm Warning, trigger "Tank1_ControlerTemp_DBW_236" bit 14
   11156: 'Tank Tank1: Heat-balancing: Motor protection supply temp. control', class Tank Alarm Warning, trigger "Tank1_ControlerTemp_DBW_236" bit 15
   11157: 'Tank Tank1: Heating: Fuse fault', class Tank Warning Archive Foaming, trigger "Tank1_ControlerTemp_DBW_236" bit 0
   11158: 'Tank Tank1: Heating: Upper limit reached', class Tank Alarm Warning, trigger "Tank1_ControlerTemp_DBW_236" bit 1
   11159: 'Tank Tank1: Heating: Lower limit reached', class Tank Alarm Warning, trigger "Tank1_ControlerTemp_DBW_236" bit 2
   11160: 'Tank Tank1: Heating: Safe shutdown reached', class Tank Alarm Warning, trigger "Tank1_ControlerTemp_DBW_236" bit 3
   11161: 'Tank Tank1: Heating: No set value specified', class Tank Alarm Warning, trigger "Tank1_ControlerTemp_DBW_236" bit 4
   11162: 'Tank Tank1: Heating:', class Tank Alarm Warning, trigger "Tank1_ControlerTemp_DBW_236" bit 5
   11163: 'Tank Tank1: Heating:', class Tank Alarm Warning, trigger "Tank1_ControlerTemp_DBW_236" bit 6
   11164: 'Tank Tank1: Heating:', class Tank Alarm Warning, trigger "Tank1_ControlerTemp_DBW_236" bit 7
   11201: 'Tank Tank2: Feed Pump: Motor Protecting switch has tripped', class Tank Alarm Warning, trigger "Tank2_FeedPump_DBW_4" bit 8
   11202: 'Tank Tank2: Feed Pump: Frequency converter fault', class Tank Alarm Warning, trigger "Tank2_FeedPump_DBW_4" bit 9
   11203: 'Tank Tank2: Feed Pump: Max.Pressure', class Tank Alarm Warning, trigger "Tank2_FeedPump_DBW_4" bit 10
   11204: 'Tank Tank2: Feed Pump: Dry run protection has tripped', class Tank Alarm Warning, trigger "Tank2_FeedPump_DBW_4" bit 11
   11205: 'Tank Tank2: Feed Pump: Wrong time entry for pause and runtime', class Tank Alarm Warning, trigger "Tank2_FeedPump_DBW_4" bit 12
   11206: 'Tank Tank2: Feed Pump: Difference pressure too high', class Tank Alarm Warning, trigger "Tank2_FeedPump_DBW_4" bit 13
   11207: 'Tank Tank2: Feed Pump: Temperature for switch-on not reached', class Tank Alarm Warning, trigger "Tank2_FeedPump_DBW_4" bit 14
   11208: 'Tank Tank2: Feed Pump: Motor protecting switch fan has tripped', class Tank Alarm Warning, trigger "Tank2_FeedPump_DBW_4" bit 15
   11209: 'Tank Tank2: Feed Pump: Filling level too low', class Tank Alarm Warning, trigger "Tank2_FeedPump_DBW_4" bit 0
   11210: 'Tank Tank2: Feed Pump: Filling selected but no barrel present', class Tank Alarm Warning, trigger "Tank2_FeedPump_DBW_4" bit 1
   11211: 'Tank Tank2: Feed Pump: No barrel present', class Tank Caution, trigger "Tank2_FeedPump_DBW_4" bit 2
   11212: 'Tank Tank2: Feed Pump:', class Tank Alarm Warning, trigger "Tank2_FeedPump_DBW_4" bit 3
   11213: 'Tank Tank2: Feed Pump:', class Tank Alarm Warning, trigger "Tank2_FeedPump_DBW_4" bit 4
   11214: 'Tank Tank2: Feed Pump:', class Tank Alarm Warning, trigger "Tank2_FeedPump_DBW_4" bit 5
   11215: 'Tank Tank2: Feed Pump:', class Tank Alarm Warning, trigger "Tank2_FeedPump_DBW_4" bit 6
   11216: 'Tank Tank2: Feed Pump:', class Tank Alarm Warning, trigger "Tank2_FeedPump_DBW_4" bit 7
   11217: 'Tank Tank2: Agitator: Motor protecting switch has tripped', class Tank Alarm Warning, trigger "Tank2_Agitator__DBW_30" bit 8
   11218: 'Tank Tank2: Agitator: Frequencny converter fault', class Tank Alarm Warning, trigger "Tank2_Agitator__DBW_30" bit 9
   11219: 'Tank Tank2: Agitator: Max drip pan filling level', class Tank Alarm Warning, trigger "Tank2_Agitator__DBW_30" bit 10
   11220: 'Tank Tank2: Agitator: Incorrect time entry for runtime or pause time', class Tank Alarm Warning, trigger "Tank2_Agitator__DBW_30" bit 11
   11221: 'Tank Tank2: Agitator:', class Tank Alarm Warning, trigger "Tank2_Agitator__DBW_30" bit 12
   11222: 'Tank Tank2: Agitator: Temperature for switch-on not reached', class Tank Alarm Warning, trigger "Tank2_Agitator__DBW_30" bit 13
   11223: 'Tank Tank2: Agitator: Fan motor protecting switch', class Tank Alarm Warning, trigger "Tank2_Agitator__DBW_30" bit 14
   11224: 'Tank Tank2: Agitator: Filling level too low', class Tank Alarm Warning, trigger "Tank2_Agitator__DBW_30" bit 15
   11225: 'Tank Tank2: Agitator:', class Tank Alarm Warning, trigger "Tank2_Agitator__DBW_30" bit 0
   11226: 'Tank Tank2: Agitator:', class Tank Alarm Warning, trigger "Tank2_Agitator__DBW_30" bit 1
   11227: 'Tank Tank2: Agitator:', class Tank Alarm Warning, trigger "Tank2_Agitator__DBW_30" bit 2
   11228: 'Tank Tank2: Agitator:', class Tank Alarm Warning, trigger "Tank2_Agitator__DBW_30" bit 3
   11229: 'Tank Tank2: Agitator:', class Tank Alarm Warning, trigger "Tank2_Agitator__DBW_30" bit 4
   11230: 'Tank Tank2: Agitator:', class Tank Alarm Warning, trigger "Tank2_Agitator__DBW_30" bit 5
   11231: 'Tank Tank2: Agitator:', class Tank Alarm Warning, trigger "Tank2_Agitator__DBW_30" bit 6
   11233: 'Tank Tank2: Filling: Min. filling level undershot', class Tank Warning Archive Foaming, trigger "Tank2_Filling_DBW_56" bit 8
   11234: 'Tank Tank2: Filling: Max. filling level exceeded', class Tank Warning Archive Foaming, trigger "Tank2_Filling_DBW_56" bit 9
   11235: 'Tank Tank2: Filling: Filling time exceeded', class Tank Alarm Warning, trigger "Tank2_Filling_DBW_56" bit 10
   11236: 'Tank Tank2: Filling: Max. drip pan filling level', class Tank Alarm Warning, trigger "Tank2_Filling_DBW_56" bit 11
   11237: 'Tank Tank2: Filling: Min. filling level in cycle', class Tank Error Filling, trigger "Tank2_Filling_DBW_56" bit 12
   11238: 'Tank Tank2: Filling: Max. filling level (with piston machines)', class Tank Error, trigger "Tank2_Filling_DBW_56" bit 13
   11239: 'Tank Tank2: Filling: Max. drip pan filling level (with piston machines)', class Tank Error Filling, trigger "Tank2_Filling_DBW_56" bit 14
   11240: 'Tank Tank2: Filling: Cable break to fill level sensor', class Tank Error Filling, trigger "Tank2_Filling_DBW_56" bit 15
   11241: 'Tank Tank2: Filling: Wrong position of fill valve', class Tank Error Filling, trigger "Tank2_Filling_DBW_56" bit 0
   11242: 'Tank Tank2: Filling: Pre-warning min. filling level', class Tank Errors Fill Archive Foaming, trigger "Tank2_Filling_DBW_56" bit 1
   11243: 'Tank Tank2: Filling:', class Tank Error Filling, trigger "Tank2_Filling_DBW_56" bit 2
   11244: 'Tank Tank2: Filling:', class Tank Error Filling, trigger "Tank2_Filling_DBW_56" bit 3
   11245: 'Tank Tank2: Filling:', class Tank Error Filling, trigger "Tank2_Filling_DBW_56" bit 4
   11246: 'Tank Tank2: Filling: Motor protection supply nucleation unit', class Tank Error Filling, trigger "Tank2_Filling_DBW_56" bit 5
   11247: 'Tank Tank2: Filling: Cable break analog value of nucleation unit', class Tank Error Filling, trigger "Tank2_Filling_DBW_56" bit 6
   11248: 'Tank Tank2: Filling: Fault from nucleation unit', class Tank Error Filling, trigger "Tank2_Filling_DBW_56" bit 7
   11249: 'Tank Tank2: Heat-balancing: Cable break to temperature sensor', class Tank Warning Archive Foaming, trigger "Tank2_ControlerTemp_DBW_238" bit 8
   11250: 'Tank Tank2: Heat-balancing: + Temperature warning', class Tank Alarm Warning, trigger "Tank2_ControlerTemp_DBW_238" bit 9
   11251: 'Tank Tank2: Heat-balancing: - Temperature warning', class Tank Alarm Warning, trigger "Tank2_ControlerTemp_DBW_238" bit 10
   11252: 'Tank Tank2: Heat-balancing: + Temperature fault', class Tank Error, trigger "Tank2_ControlerTemp_DBW_238" bit 11
   11253: 'Tank Tank2: Heat-balancing: - Temperature fault', class Tank Error, trigger "Tank2_ControlerTemp_DBW_238" bit 12
   11254: 'Tank Tank2: Heat-balancing:Controller at limit', class Tank Alarm Warning, trigger "Tank2_ControlerTemp_DBW_238" bit 13
   11255: 'Tank Tank2: Heat-balancing:', class Tank Alarm Warning, trigger "Tank2_ControlerTemp_DBW_238" bit 14
   11256: 'Tank Tank2: Heat-balancing: Motor protection supply temp. control', class Tank Alarm Warning, trigger "Tank2_ControlerTemp_DBW_238" bit 15
   11257: 'Tank Tank2: Heating: Fuse fault', class Tank Warning Archive Foaming, trigger "Tank2_ControlerTemp_DBW_238" bit 0
   11258: 'Tank Tank2: Heating: Upper limit reached', class Tank Alarm Warning, trigger "Tank2_ControlerTemp_DBW_238" bit 1
   11259: 'Tank Tank2: Heating: Lower limit reached', class Tank Alarm Warning, trigger "Tank2_ControlerTemp_DBW_238" bit 2
   11260: 'Tank Tank2: Heating: Safe shutdown reached', class Tank Alarm Warning, trigger "Tank2_ControlerTemp_DBW_238" bit 3
   11261: 'Tank Tank2: Heating: No set value specified', class Tank Alarm Warning, trigger "Tank2_ControlerTemp_DBW_238" bit 4
   11262: 'Tank Tank2: Heating:', class Tank Alarm Warning, trigger "Tank2_ControlerTemp_DBW_238" bit 5
   11263: 'Tank Tank2: Heating:', class Tank Alarm Warning, trigger "Tank2_ControlerTemp_DBW_238" bit 6
   11264: 'Tank Tank2: Heating:', class Tank Alarm Warning, trigger "Tank2_ControlerTemp_DBW_238" bit 7
   11381: 'Tank Tank1: Pentane: Pre alarm for pentane (20%)', class Tank Alarm Warning, trigger "Tank1_Pentan_DBW_496" bit 8
   11382: 'Tank Tank1: Pentane: Pre alarm nitrogen at the tank low', class Tank Alarm Warning, trigger "Tank1_Pentan_DBW_496" bit 9
   11383: 'Tank Tank1: Pentane: Nitrogen pressure at the tank low', class Tank Alarm Warning, trigger "Tank1_Pentan_DBW_496" bit 10
   11384: 'Tank Tank1: Pentane: Nitrogen supply low', class Tank Alarm Warning, trigger "Tank1_Pentan_DBW_496" bit 11
   11385: 'Tank Tank1: Pentane: Exhaust system not ready', class Tank Alarm Warning, trigger "Tank1_Pentan_DBW_496" bit 12
   11386: 'Tank Tank1: Pentane: Supply pump not running', class Tank Alarm Warning, trigger "Tank1_Pentan_DBW_496" bit 13
   11387: 'Tank Tank1: Pentane: Pertamix not ready', class Tank Caution, trigger "Tank1_Pentan_DBW_496" bit 14
   11388: 'Tank Tank1: Pentane: Emergency stop from pertamix exists', class Tank Alarm Warning, trigger "Tank1_Pentan_DBW_496" bit 15
   11389: 'Tank Tank1: Pentane: Filling valve 1 not close', class Tank Alarm Warning, trigger "Tank1_Pentan_DBW_496" bit 0
   11390: 'Tank Tank1: Pentane: Filling valve 2 not close', class Tank Alarm Warning, trigger "Tank1_Pentan_DBW_496" bit 1
   11391: 'Tank Tank1: Pentane: No start signal from the scales', class Tank Alarm Warning, trigger "Tank1_Pentan_DBW_496" bit 2
   11392: 'Tank Tank1: Pentane: No source (Poly or Pentane) selected', class Tank Alarm Warning, trigger "Tank1_Pentan_DBW_496" bit 3
   11393: 'Tank Tank1: Pentane:', class Tank Alarm Warning, trigger "Tank1_Pentan_DBW_496" bit 4
   11394: 'Tank Tank1: Pentane:', class Tank Alarm Warning, trigger "Tank1_Pentan_DBW_496" bit 5
   11395: 'Tank Tank1: Pentane:', class Tank Alarm Warning, trigger "Tank1_Pentan_DBW_496" bit 6
   11396: 'Tank Tank1: Pentane:', class Tank Alarm Warning, trigger "Tank1_Pentan_DBW_496" bit 7
   713: 'Tank Tank1:', class Tank Alarm Warning, trigger "Interface_Container_DBW_520" bit 4
   714: 'Tank Tank1:', class Tank Alarm Warning, trigger "Interface_Container_DBW_520" bit 5
   715: 'Tank Tank1:', class Tank Alarm Warning, trigger "Interface_Container_DBW_520" bit 6
   716: 'Tank Tank1:', class Tank Alarm Warning, trigger "Interface_Container_DBW_520" bit 7
   12101: 'Pump1: FeedPump: motor protecting switch has tripped', class Pump Warning Alarm, trigger "Pump1_FeedPump_DBW_2" bit 8
   12102: 'Pump1: FeedPump: frequency converter fault', class Pump Warning Alarm, trigger "Pump1_FeedPump_DBW_2" bit 9